TYPE "Table Row Data"
   STRUCT
      address : UInt;
      ordered : Bool;
      pbSelection : Struct
         actuate : Bool;
         animate : USInt;
      END_STRUCT;
      rtBackground : Struct
         animate : USInt;
      END_STRUCT;
      tfDropZone : Struct
         animate : USInt;
         value : WString[20];
      END_STRUCT;
      tfLine : Struct
         animate : USInt;
         value : WString[20];
      END_STRUCT;
      tfPartNumber : Struct
         animateDL : USInt;
         animateSL : USInt;
         value : WString[40];
      END_STRUCT;
      tfTime : Struct
         animate : USInt;
         value : WString[20];
      END_STRUCT;
   END_STRUCT;
END_TYPE

TYPE "Station Assignment: Button Details Data"
   STRUCT
      alloted : Struct
         animate : USInt;
         value : WString[10];
      END_STRUCT;
      critical : Struct
         animate : USInt;
         value : WString[10];
      END_STRUCT;
      label : Struct
         animate : USInt;
         value : WString[2];
      END_STRUCT;
      partNumber : Struct
         animate : USInt;
         value : WString[40];
      END_STRUCT;
      select : Struct
         actuate : Bool;
         animate : USInt;
      END_STRUCT;
   END_STRUCT;
END_TYPE

(* ===== HMI "HMI_RT_1" =====
system functions are stored by id; their names below are inferred from use
connection "HMI_Connection_2": ETHERNET, S7_1500_OMS

HMI tags "Default tag table"
   "Clock_Byte" : Byte = PLC Clock_Byte AT %MB0, 100 ms
   "HMI_screenNumber" : Int = PLC HMI.screenNumber AT %DB1.DBW0, 100 ms
   "HMI_barcode" : Barcode Screen = PLC HMI.barcode AT %DB1.DBW0, 100 ms
   "HMI_partCall_row{0}" : Table Row = PLC HMI.partCall.row[0], 100 ms
   "HMI_partCall_row{1}" : Table Row = PLC HMI.partCall.row[1], 100 ms
   "HMI_partCall_row{2}" : Table Row = PLC HMI.partCall.row[2], 100 ms
   "HMI_partCall_row{3}" : Table Row = PLC HMI.partCall.row[3], 100 ms
   "HMI_partCall_row{4}" : Table Row = PLC HMI.partCall.row[4], 100 ms
   "HMI_partCall_row{5}" : Table Row = PLC HMI.partCall.row[5], 100 ms
   "HMI_partCall_row{6}" : Table Row = PLC HMI.partCall.row[6], 100 ms
   "HMI_partCall_row{7}" : Table Row = PLC HMI.partCall.row[7], 100 ms
   "HMI_partCall_row{8}" : Table Row = PLC HMI.partCall.row[8], 100 ms
   "HMI_partCall_row{9}" : Table Row = PLC HMI.partCall.row[9], 100 ms
   "HMI_partCall_row{10}" : Table Row = PLC HMI.partCall.row[10], 100 ms
   "HMI_settings_stations_selectBtns{0}" : PB Data: Text Label = PLC HMI.settings.stations.selectBtns[0], 100 ms
   "HMI_settings_stations_selectBtns{1}" : PB Data: Text Label = PLC HMI.settings.stations.selectBtns[1], 100 ms
   "HMI_settings_stations_selectBtns{2}" : PB Data: Text Label = PLC HMI.settings.stations.selectBtns[2], 100 ms
   "HMI_settings_stations_selectBtns{3}" : PB Data: Text Label = PLC HMI.settings.stations.selectBtns[3], 100 ms
   "HMI_settings_stations_selectBtns{4}" : PB Data: Text Label = PLC HMI.settings.stations.selectBtns[4], 100 ms
   "HMI_settings_stations_selectBtns{5}" : PB Data: Text Label = PLC HMI.settings.stations.selectBtns[5], 100 ms
   "HMI_settings_stations_selectBtns{6}" : PB Data: Text Label = PLC HMI.settings.stations.selectBtns[6], 100 ms
   "HMI_settings_stations_selectBtns{7}" : PB Data: Text Label = PLC HMI.settings.stations.selectBtns[7], 100 ms
   "HMI_settings_stations_selectBtns{8}" : PB Data: Text Label = PLC HMI.settings.stations.selectBtns[8], 100 ms
   "HMI_settings_stations_selectBtns{9}" : PB Data: Text Label = PLC HMI.settings.stations.selectBtns[9], 100 ms
   "HMI_settings_stations_selectBtns{10}" : PB Data: Text Label = PLC HMI.settings.stations.selectBtns[10], 100 ms
   "HMI_settings_stations_selectBtns{11}" : PB Data: Text Label = PLC HMI.settings.stations.selectBtns[11], 100 ms
   "HMI_settings_kp8_buttons{0}" : PB Data: Text Label = PLC HMI.settings.kp8.buttons[0], 100 ms
   "HMI_settings_kp8_buttons{7}" : PB Data: Text Label = PLC HMI.settings.kp8.buttons[7], 100 ms
   "HMI_settings_kp8_buttons{3}" : PB Data: Text Label = PLC HMI.settings.kp8.buttons[3], 100 ms
   "HMI_settings_kp8_buttons{6}" : PB Data: Text Label = PLC HMI.settings.kp8.buttons[6], 100 ms
   "HMI_settings_kp8_buttons{2}" : PB Data: Text Label = PLC HMI.settings.kp8.buttons[2], 100 ms
   "HMI_settings_kp8_buttons{5}" : PB Data: Text Label = PLC HMI.settings.kp8.buttons[5], 100 ms
   "HMI_settings_kp8_buttons{1}" : PB Data: Text Label = PLC HMI.settings.kp8.buttons[1], 100 ms
   "HMI_settings_kp8_buttons{4}" : PB Data: Text Label = PLC HMI.settings.kp8.buttons[4], 100 ms
   "HMI_settings_stations_selCount" : Int = PLC HMI.settings.stations.selCount, 100 ms
   "HMI_settings_viewingStation_btns{0}" : Station Assignment: Button Details = PLC HMI.settings.viewingStation.btns[0], 100 ms
   "HMI_settings_viewingStation_btns{1}" : Station Assignment: Button Details = PLC HMI.settings.viewingStation.btns[1], 100 ms
   "HMI_settings_viewingStation_btns{2}" : Station Assignment: Button Details = PLC HMI.settings.viewingStation.btns[2], 100 ms
   "HMI_settings_viewingStation_btns{3}" : Station Assignment: Button Details = PLC HMI.settings.viewingStation.btns[3], 100 ms
   "HMI_settings_viewingStation_btns{4}" : Station Assignment: Button Details = PLC HMI.settings.viewingStation.btns[4], 100 ms
   "HMI_settings_viewingStation_btns{5}" : Station Assignment: Button Details = PLC HMI.settings.viewingStation.btns[5], 100 ms
   "HMI_settings_viewingStation_previous" : PB Data: Graphic/Text List = PLC HMI.settings.viewingStation.previous, 100 ms
   "HMI_settings_viewingStation_next" : PB Data: Graphic/Text List = PLC HMI.settings.viewingStation.next, 100 ms
   "HMI_settings_stations_selectAll" : PB Data: Text Label = PLC HMI.settings.stations.selectAll, 100 ms
   "HMI_settings_partNumber_assign" : PB Data: Text Label = PLC HMI.settings.partNumber.assign, 100 ms
   "HMI_settings_partNumber_ioField" : IO Field Data: Part Number = PLC HMI.settings.partNumber.ioField, 100 ms
   "HMI_settings_alotted_assign" : PB Data: Text Label = PLC HMI.settings.alotted.assign, 100 ms
   "HMI_settings_alotted_ioField" : IO Field Data: Timers = PLC HMI.settings.alotted.ioField, 100 ms
   "HMI_settings_critical_assign" : PB Data: Text Label = PLC HMI.settings.critical.assign, 100 ms
   "HMI_settings_critical_ioField" : IO Field Data: Timers = PLC HMI.settings.critical.ioField, 100 ms
   "HMI_settings_kp8_selectButtons" : PB Data: Text Label = PLC HMI.settings.kp8.selectButtons, 100 ms
   "HMI_settings_viewingStation_dzData" : Drop Zone Data = PLC HMI.settings.viewingStation.dzData, 100 ms
   "HMI_settings_viewingStation_lineData" : Line Label Data = PLC HMI.settings.viewingStation.lineData, 100 ms
   "HMI_settings_stations_prevGroup" : PB Data: Graphic/Text List = PLC HMI.settings.stations.prevGroup, 100 ms
   "HMI_settings_stations_nextGroup" : PB Data: Graphic/Text List = PLC HMI.settings.stations.nextGroup, 100 ms
   "HMI_settings_viewingStation_name" : WString[20] = PLC HMI.settings.viewingStation.name, 100 ms
   "HMI_tableNav_top" : PB Data: Graphic/Text List = PLC HMI.tableNav.top, 100 ms
   "HMI_tableNav_pageUp" : PB Data: Graphic/Text List = PLC HMI.tableNav.pageUp, 100 ms
   "HMI_tableNav_lineUp" : PB Data: Graphic/Text List = PLC HMI.tableNav.lineUp, 100 ms
   "HMI_tableNav_lineDown" : PB Data: Graphic/Text List = PLC HMI.tableNav.lineDown, 100 ms
   "HMI_tableNav_pageDown" : PB Data: Graphic/Text List = PLC HMI.tableNav.pageDown, 100 ms
   "HMI_tableNav_bottom" : PB Data: Graphic/Text List = PLC HMI.tableNav.bottom, 100 ms
   "HMI_simStations_stations{0}" : Station Sim Data = PLC HMI.simStations.me[0] AT %DB1.DBX0.0, 100 ms
   "HMI_simStations_me{1}" : Station Sim Data = PLC HMI.simStations.me[1], 100 ms
   "HMI_simStations_me{2}" : Station Sim Data = PLC HMI.simStations.me[2], 100 ms
   "HMI_simStations_me{3}" : Station Sim Data = PLC HMI.simStations.me[3], 100 ms
   "HMI_simStations_me{4}" : Station Sim Data = PLC HMI.simStations.me[4], 100 ms
   "HMI_simStations_me{5}" : Station Sim Data = PLC HMI.simStations.me[5], 100 ms
   "HMI_simStations_me{6}" : Station Sim Data = PLC HMI.simStations.me[6], 100 ms
   "HMI_simStations_me{7}" : Station Sim Data = PLC HMI.simStations.me[7], 100 ms
   "HMI_simStations_me{8}" : Station Sim Data = PLC HMI.simStations.me[8], 100 ms
   "HMI_simStations_me{9}" : Station Sim Data = PLC HMI.simStations.me[9], 100 ms
   "HMI_simStations_me{10}" : Station Sim Data = PLC HMI.simStations.me[10], 100 ms
   "HMI_simStations_me{11}" : Station Sim Data = PLC HMI.simStations.me[11], 100 ms
   "HMI_simStations_up" : PB Data: Graphic/Text List = PLC HMI.simStations.up, 100 ms
   "HMI_simStations_down" : PB Data: Graphic/Text List = PLC HMI.simStations.down, 100 ms
   "Log Flag" : Int = PLC "Log Buffer".logFlag AT %DB1.DBW0, 100 ms
      on ChangeValue: function_abcfba0d("Log Buffer_partReq_me{0}_address"); function_abcfba0d("Log Buffer_partReq_me{0}_timeStamp"); function_abcfba0d("Log Buffer_partReq_me{0}_reqType")
   "Log Buffer_partReq_me{0}_address" : Int = PLC "Log Buffer".partReq.me[0].address, 100 ms
   "Log Buffer_partReq_me{0}_timeStamp" : DTL = PLC "Log Buffer".partReq.me[0].timeStamp, 100 ms
   "Log Buffer_partReq_me{0}_reqType" : Int = PLC "Log Buffer".partReq.me[0].reqType, 100 ms
   "HMI_networkHealth_pnioDevices{1}" : PB Data: Text Label = PLC HMI.networkHealth.pnioDevices[1], 100 ms
   "HMI_networkHealth_pnioDevices{2}" : PB Data: Text Label = PLC HMI.networkHealth.pnioDevices[2], 1 s
   "HMI_networkHealth_pnioDevices{3}" : PB Data: Text Label = PLC HMI.networkHealth.pnioDevices[3], 1 s
   "HMI_networkHealth_pnioDevices{4}" : PB Data: Text Label = PLC HMI.networkHealth.pnioDevices[4], 1 s
   "HMI_networkHealth_pnioDevices{5}" : PB Data: Text Label = PLC HMI.networkHealth.pnioDevices[5], 1 s
   "HMI_networkHealth_pnioDevices{6}" : PB Data: Text Label = PLC HMI.networkHealth.pnioDevices[6], 1 s
   "HMI_networkHealth_pnioDevices{7}" : PB Data: Text Label = PLC HMI.networkHealth.pnioDevices[7], 1 s
   "HMI_networkHealth_pnioDevices{8}" : PB Data: Text Label = PLC HMI.networkHealth.pnioDevices[8], 1 s
   "HMI_networkHealth_pnioDevices{9}" : PB Data: Text Label = PLC HMI.networkHealth.pnioDevices[9], 1 s
   "HMI_networkHealth_pnioDevices{10}" : PB Data: Text Label = PLC HMI.networkHealth.pnioDevices[10], 1 s
   "HMI_networkHealth_pnioDevices{11}" : PB Data: Text Label = PLC HMI.networkHealth.pnioDevices[11], 1 s
   "HMI_networkHealth_pnioDevices{12}" : PB Data: Text Label = PLC HMI.networkHealth.pnioDevices[12], 1 s
   "HMI_networkHealth_pnioDevices{13}" : PB Data: Text Label = PLC HMI.networkHealth.pnioDevices[13], 1 s
   "HMI_networkHealth_pnioDevices{16}" : PB Data: Text Label = PLC HMI.networkHealth.pnioDevices[16], 1 s
   "HMI_networkHealth_pnioDevices{14}" : PB Data: Text Label = PLC HMI.networkHealth.pnioDevices[14], 1 s
   "HMI_networkHealth_pnioDevices{15}" : PB Data: Text Label = PLC HMI.networkHealth.pnioDevices[15], 1 s
   "HMI_networkHealth_pnioDevices{17}" : PB Data: Text Label = PLC HMI.networkHealth.pnioDevices[17], 1 s
   "HMI_networkHealth_pnioDevices{18}" : PB Data: Text Label = PLC HMI.networkHealth.pnioDevices[18], 1 s
   "HMI_networkHealth_pnioDevices{19}" : PB Data: Text Label = PLC HMI.networkHealth.pnioDevices[19], 1 s
   "HMI_networkHealth_pnioDevices{20}" : PB Data: Text Label = PLC HMI.networkHealth.pnioDevices[20], 1 s
   "HMI_networkHealth_pnioDevices{21}" : PB Data: Text Label = PLC HMI.networkHealth.pnioDevices[21], 1 s
   "HMI_networkHealth_pnioDevices{22}" : PB Data: Text Label = PLC HMI.networkHealth.pnioDevices[22], 1 s
   "HMI_networkHealth_pnioDevices{31}" : PB Data: Text Label = PLC HMI.networkHealth.pnioDevices[31], 1 s
   "HMI_networkHealth_pnioDevices{32}" : PB Data: Text Label = PLC HMI.networkHealth.pnioDevices[32], 1 s
   "HMI_networkHealth_pnioDevices{29}" : PB Data: Text Label = PLC HMI.networkHealth.pnioDevices[29], 1 s
   "HMI_networkHealth_pnioDevices{30}" : PB Data: Text Label = PLC HMI.networkHealth.pnioDevices[30], 1 s
   "HMI_networkHealth_pnioDevices{27}" : PB Data: Text Label = PLC HMI.networkHealth.pnioDevices[27], 1 s
   "HMI_networkHealth_pnioDevices{28}" : PB Data: Text Label = PLC HMI.networkHealth.pnioDevices[28], 1 s
   "HMI_networkHealth_pnioDevices{23}" : PB Data: Text Label = PLC HMI.networkHealth.pnioDevices[23], 1 s
   "HMI_networkHealth_pnioDevices{24}" : PB Data: Text Label = PLC HMI.networkHealth.pnioDevices[24], 1 s
   "HMI_networkHealth_pnioDevices{25}" : PB Data: Text Label = PLC HMI.networkHealth.pnioDevices[25], 1 s
   "HMI_networkHealth_pnioDevices{26}" : PB Data: Text Label = PLC HMI.networkHealth.pnioDevices[26], 1 s
   "HMI_networkHealth_pnioDevices{33}" : PB Data: Text Label = PLC HMI.networkHealth.pnioDevices[33], 1 s
   "HMI_networkHealth_pnioDevices{34}" : PB Data: Text Label = PLC HMI.networkHealth.pnioDevices[34], 1 s
   "HMI_networkHealth_pnioDevices{35}" : PB Data: Text Label = PLC HMI.networkHealth.pnioDevices[35], 1 s
   "HMI_networkHealth_pnioDevices{36}" : PB Data: Text Label = PLC HMI.networkHealth.pnioDevices[36], 1 s
   "HMI_networkHealth_pnioDevices{37}" : PB Data: Text Label = PLC HMI.networkHealth.pnioDevices[37], 1 s
   "HMI_networkHealth_pnioDevices{38}" : PB Data: Text Label = PLC HMI.networkHealth.pnioDevices[38], 1 s
   "HMI_networkHealth_pnioDevices{39}" : PB Data: Text Label = PLC HMI.networkHealth.pnioDevices[39], 1 s
   "HMI_networkHealth_pnioDevices{40}" : PB Data: Text Label = PLC HMI.networkHealth.pnioDevices[40], 1 s
   "HMI_networkHealth_pnioDevices{41}" : PB Data: Text Label = PLC HMI.networkHealth.pnioDevices[41], 1 s
   "HMI_networkHealth_pnioDevices{42}" : PB Data: Text Label = PLC HMI.networkHealth.pnioDevices[42], 1 s
   "HMI_networkHealth_pnioDevices{43}" : PB Data: Text Label = PLC HMI.networkHealth.pnioDevices[43], 1 s
   "HMI_networkHealth_pnioDevices{44}" : PB Data: Text Label = PLC HMI.networkHealth.pnioDevices[44], 1 s
   "HMI_networkHealth_pnioDevices{45}" : PB Data: Text Label = PLC HMI.networkHealth.pnioDevices[45], 1 s
   "HMI_networkHealth_pnioDevices{46}" : PB Data: Text Label = PLC HMI.networkHealth.pnioDevices[46], 1 s
   "HMI_networkHealth_pnioDevices{47}" : PB Data: Text Label = PLC HMI.networkHealth.pnioDevices[47], 1 s
   "HMI_networkHealth_pnioDevices{48}" : PB Data: Text Label = PLC HMI.networkHealth.pnioDevices[48], 1 s
   "HMI_networkHealth_et200spPopUp" : Station: ET200SP Comm Debug Data = PLC HMI.networkHealth.et200spPopUp, 1 s
   "HMI_networkHealth_kp8PopUp" : Station: KP8 Comm Debug Data = PLC HMI.networkHealth.kp8PopUp, 1 s
   "HMI_networkHealth_selectedDevice" : Int = PLC HMI.networkHealth.selectedDevice, 1 s
   "EMP IDB_stations_me{0}_partNumbers{0}" : WString[40] = PLC "EMP IDB".stations.me[0].partNumbers[0], 1 s
   "EMP IDB_stations_me{0}_partNumbers{1}" : WString[40] = PLC "EMP IDB".stations.me[0].partNumbers[1], 1 s
   "EMP IDB_stations_me{0}_partNumbers{2}" : WString[40] = PLC "EMP IDB".stations.me[0].partNumbers[2], 1 s
   "EMP IDB_stations_me{0}_partNumbers{3}" : WString[40] = PLC "EMP IDB".stations.me[0].partNumbers[3], 1 s
   "EMP IDB_stations_me{0}_partNumbers{4}" : WString[40] = PLC "EMP IDB".stations.me[0].partNumbers[4], 1 s
   "EMP IDB_stations_me{0}_partNumbers{5}" : WString[40] = PLC "EMP IDB".stations.me[0].partNumbers[5], 1 s
   "EMP IDB_stations_me{0}_partNumbers{6}" : WString[40] = PLC "EMP IDB".stations.me[0].partNumbers[6], 1 s
   "EMP IDB_stations_me{0}_partNumbers{7}" : WString[40] = PLC "EMP IDB".stations.me[0].partNumbers[7], 1 s
   "EMP IDB_stations_me{1}_partNumbers{0}" : WString[40] = PLC "EMP IDB".stations.me[1].partNumbers[0], 1 s
   "EMP IDB_stations_me{1}_partNumbers{1}" : WString[40] = PLC "EMP IDB".stations.me[1].partNumbers[1], 1 s
   "EMP IDB_stations_me{1}_partNumbers{2}" : WString[40] = PLC "EMP IDB".stations.me[1].partNumbers[2], 1 s
   "EMP IDB_stations_me{1}_partNumbers{3}" : WString[40] = PLC "EMP IDB".stations.me[1].partNumbers[3], 1 s
   "EMP IDB_stations_me{1}_partNumbers{4}" : WString[40] = PLC "EMP IDB".stations.me[1].partNumbers[4], 1 s
   "EMP IDB_stations_me{1}_partNumbers{5}" : WString[40] = PLC "EMP IDB".stations.me[1].partNumbers[5], 1 s
   "EMP IDB_stations_me{1}_partNumbers{6}" : WString[40] = PLC "EMP IDB".stations.me[1].partNumbers[6], 1 s
   "EMP IDB_stations_me{1}_partNumbers{7}" : WString[40] = PLC "EMP IDB".stations.me[1].partNumbers[7], 1 s
   "EMP IDB_stations_me{2}_partNumbers{0}" : WString[40] = PLC "EMP IDB".stations.me[2].partNumbers[0], 1 s
   "EMP IDB_stations_me{2}_partNumbers{1}" : WString[40] = PLC "EMP IDB".stations.me[2].partNumbers[1], 1 s
   "EMP IDB_stations_me{2}_partNumbers{2}" : WString[40] = PLC "EMP IDB".stations.me[2].partNumbers[2], 1 s
   "EMP IDB_stations_me{2}_partNumbers{3}" : WString[40] = PLC "EMP IDB".stations.me[2].partNumbers[3], 1 s
   "EMP IDB_stations_me{2}_partNumbers{4}" : WString[40] = PLC "EMP IDB".stations.me[2].partNumbers[4], 1 s
   "EMP IDB_stations_me{2}_partNumbers{5}" : WString[40] = PLC "EMP IDB".stations.me[2].partNumbers[5], 1 s
   "EMP IDB_stations_me{2}_partNumbers{6}" : WString[40] = PLC "EMP IDB".stations.me[2].partNumbers[6], 1 s
   "EMP IDB_stations_me{2}_partNumbers{7}" : WString[40] = PLC "EMP IDB".stations.me[2].partNumbers[7], 1 s
   "EMP IDB_stations_me{3}_partOrdered{0}" : Bool = PLC "EMP IDB".stations.me[3].partOrdered[0], 1 s
   "EMP IDB_stations_me{3}_partOrdered{1}" : Bool = PLC "EMP IDB".stations.me[3].partOrdered[1], 1 s
   "EMP IDB_stations_me{3}_partOrdered{2}" : Bool = PLC "EMP IDB".stations.me[3].partOrdered[2], 1 s
   "EMP IDB_stations_me{3}_partOrdered{3}" : Bool = PLC "EMP IDB".stations.me[3].partOrdered[3], 1 s
   "EMP IDB_stations_me{3}_partOrdered{4}" : Bool = PLC "EMP IDB".stations.me[3].partOrdered[4], 1 s
   "EMP IDB_stations_me{3}_partOrdered{5}" : Bool = PLC "EMP IDB".stations.me[3].partOrdered[5], 1 s
   "EMP IDB_stations_me{3}_partOrdered{6}" : Bool = PLC "EMP IDB".stations.me[3].partOrdered[6], 1 s
   "EMP IDB_stations_me{3}_partOrdered{7}" : Bool = PLC "EMP IDB".stations.me[3].partOrdered[7], 1 s
   "EMP IDB_stations_me{4}_partNumbers{0}" : WString[40] = PLC "EMP IDB".stations.me[4].partNumbers[0], 1 s
   "EMP IDB_stations_me{4}_partNumbers{1}" : WString[40] = PLC "EMP IDB".stations.me[4].partNumbers[1], 1 s
   "EMP IDB_stations_me{4}_partNumbers{2}" : WString[40] = PLC "EMP IDB".stations.me[4].partNumbers[2], 1 s
   "EMP IDB_stations_me{4}_partNumbers{3}" : WString[40] = PLC "EMP IDB".stations.me[4].partNumbers[3], 1 s
   "EMP IDB_stations_me{4}_partNumbers{4}" : WString[40] = PLC "EMP IDB".stations.me[4].partNumbers[4], 1 s
   "EMP IDB_stations_me{4}_partNumbers{5}" : WString[40] = PLC "EMP IDB".stations.me[4].partNumbers[5], 1 s
   "EMP IDB_stations_me{4}_partNumbers{6}" : WString[40] = PLC "EMP IDB".stations.me[4].partNumbers[6], 1 s
   "EMP IDB_stations_me{4}_partNumbers{7}" : WString[40] = PLC "EMP IDB".stations.me[4].partNumbers[7], 1 s
   "EMP IDB_stations_me{5}_partNumbers{0}" : WString[40] = PLC "EMP IDB".stations.me[5].partNumbers[0], 1 s
   "EMP IDB_stations_me{5}_partNumbers{1}" : WString[40] = PLC "EMP IDB".stations.me[5].partNumbers[1], 1 s
   "EMP IDB_stations_me{5}_partNumbers{2}" : WString[40] = PLC "EMP IDB".stations.me[5].partNumbers[2], 1 s
   "EMP IDB_stations_me{5}_partNumbers{3}" : WString[40] = PLC "EMP IDB".stations.me[5].partNumbers[3], 1 s
   "EMP IDB_stations_me{5}_partNumbers{4}" : WString[40] = PLC "EMP IDB".stations.me[5].partNumbers[4], 1 s
   "EMP IDB_stations_me{5}_partNumbers{5}" : WString[40] = PLC "EMP IDB".stations.me[5].partNumbers[5], 1 s
   "EMP IDB_stations_me{5}_partNumbers{6}" : WString[40] = PLC "EMP IDB".stations.me[5].partNumbers[6], 1 s
   "EMP IDB_stations_me{5}_partNumbers{7}" : WString[40] = PLC "EMP IDB".stations.me[5].partNumbers[7], 1 s
   "EMP IDB_stations_me{6}_partNumbers{0}" : WString[40] = PLC "EMP IDB".stations.me[6].partNumbers[0], 1 s
   "EMP IDB_stations_me{6}_partNumbers{1}" : WString[40] = PLC "EMP IDB".stations.me[6].partNumbers[1], 1 s
   "EMP IDB_stations_me{6}_partNumbers{2}" : WString[40] = PLC "EMP IDB".stations.me[6].partNumbers[2], 1 s
   "EMP IDB_stations_me{6}_partNumbers{3}" : WString[40] = PLC "EMP IDB".stations.me[6].partNumbers[3], 1 s
   "EMP IDB_stations_me{6}_partNumbers{4}" : WString[40] = PLC "EMP IDB".stations.me[6].partNumbers[4], 1 s
   "EMP IDB_stations_me{6}_partNumbers{5}" : WString[40] = PLC "EMP IDB".stations.me[6].partNumbers[5], 1 s
   "EMP IDB_stations_me{6}_partNumbers{6}" : WString[40] = PLC "EMP IDB".stations.me[6].partNumbers[6], 1 s
   "EMP IDB_stations_me{6}_partNumbers{7}" : WString[40] = PLC "EMP IDB".stations.me[6].partNumbers[7], 1 s
   "EMP IDB_stations_me{7}_partNumbers{0}" : WString[40] = PLC "EMP IDB".stations.me[7].partNumbers[0], 1 s
   "EMP IDB_stations_me{7}_partNumbers{1}" : WString[40] = PLC "EMP IDB".stations.me[7].partNumbers[1], 1 s
   "EMP IDB_stations_me{7}_partNumbers{2}" : WString[40] = PLC "EMP IDB".stations.me[7].partNumbers[2], 1 s
   "EMP IDB_stations_me{7}_partNumbers{3}" : WString[40] = PLC "EMP IDB".stations.me[7].partNumbers[3], 1 s
   "EMP IDB_stations_me{7}_partNumbers{4}" : WString[40] = PLC "EMP IDB".stations.me[7].partNumbers[4], 1 s
   "EMP IDB_stations_me{7}_partNumbers{5}" : WString[40] = PLC "EMP IDB".stations.me[7].partNumbers[5], 1 s
   "EMP IDB_stations_me{7}_partNumbers{6}" : WString[40] = PLC "EMP IDB".stations.me[7].partNumbers[6], 1 s
   "EMP IDB_stations_me{7}_partNumbers{7}" : WString[40] = PLC "EMP IDB".stations.me[7].partNumbers[7], 1 s
   "EMP IDB_stations_me{8}_partNumbers{0}" : WString[40] = PLC "EMP IDB".stations.me[8].partNumbers[0], 1 s
   "EMP IDB_stations_me{8}_partNumbers{1}" : WString[40] = PLC "EMP IDB".stations.me[8].partNumbers[1], 1 s
   "EMP IDB_stations_me{8}_partNumbers{2}" : WString[40] = PLC "EMP IDB".stations.me[8].partNumbers[2], 1 s
   "EMP IDB_stations_me{8}_partNumbers{3}" : WString[40] = PLC "EMP IDB".stations.me[8].partNumbers[3], 1 s
   "EMP IDB_stations_me{8}_partNumbers{4}" : WString[40] = PLC "EMP IDB".stations.me[8].partNumbers[4], 1 s
   "EMP IDB_stations_me{8}_partNumbers{5}" : WString[40] = PLC "EMP IDB".stations.me[8].partNumbers[5], 1 s
   "EMP IDB_stations_me{8}_partNumbers{6}" : WString[40] = PLC "EMP IDB".stations.me[8].partNumbers[6], 1 s
   "EMP IDB_stations_me{8}_partNumbers{7}" : WString[40] = PLC "EMP IDB".stations.me[8].partNumbers[7], 1 s
   "EMP IDB_stations_me{9}_partNumbers{0}" : WString[40] = PLC "EMP IDB".stations.me[9].partNumbers[0], 1 s
   "EMP IDB_stations_me{9}_partNumbers{1}" : WString[40] = PLC "EMP IDB".stations.me[9].partNumbers[1], 1 s
   "EMP IDB_stations_me{9}_partNumbers{2}" : WString[40] = PLC "EMP IDB".stations.me[9].partNumbers[2], 1 s
   "EMP IDB_stations_me{9}_partNumbers{3}" : WString[40] = PLC "EMP IDB".stations.me[9].partNumbers[3], 1 s
   "EMP IDB_stations_me{9}_partNumbers{4}" : WString[40] = PLC "EMP IDB".stations.me[9].partNumbers[4], 1 s
   "EMP IDB_stations_me{9}_partNumbers{5}" : WString[40] = PLC "EMP IDB".stations.me[9].partNumbers[5], 1 s
   "EMP IDB_stations_me{9}_partNumbers{6}" : WString[40] = PLC "EMP IDB".stations.me[9].partNumbers[6], 1 s
   "EMP IDB_stations_me{9}_partNumbers{7}" : WString[40] = PLC "EMP IDB".stations.me[9].partNumbers[7], 1 s
   "EMP IDB_stations_me{10}_partNumbers{0}" : WString[40] = PLC "EMP IDB".stations.me[10].partNumbers[0], 1 s
   "EMP IDB_stations_me{10}_partNumbers{1}" : WString[40] = PLC "EMP IDB".stations.me[10].partNumbers[1], 1 s
   "EMP IDB_stations_me{10}_partNumbers{2}" : WString[40] = PLC "EMP IDB".stations.me[10].partNumbers[2], 1 s
   "EMP IDB_stations_me{10}_partNumbers{3}" : WString[40] = PLC "EMP IDB".stations.me[10].partNumbers[3], 1 s
   "EMP IDB_stations_me{10}_partNumbers{4}" : WString[40] = PLC "EMP IDB".stations.me[10].partNumbers[4], 1 s
   "EMP IDB_stations_me{10}_partNumbers{5}" : WString[40] = PLC "EMP IDB".stations.me[10].partNumbers[5], 1 s
   "EMP IDB_stations_me{10}_partNumbers{6}" : WString[40] = PLC "EMP IDB".stations.me[10].partNumbers[6], 1 s
   "EMP IDB_stations_me{10}_partNumbers{7}" : WString[40] = PLC "EMP IDB".stations.me[10].partNumbers[7], 1 s
   "EMP IDB_stations_me{11}_partNumbers{0}" : WString[40] = PLC "EMP IDB".stations.me[11].partNumbers[0], 1 s
   "EMP IDB_stations_me{11}_partNumbers{1}" : WString[40] = PLC "EMP IDB".stations.me[11].partNumbers[1], 1 s
   "EMP IDB_stations_me{11}_partNumbers{2}" : WString[40] = PLC "EMP IDB".stations.me[11].partNumbers[2], 1 s
   "EMP IDB_stations_me{11}_partNumbers{3}" : WString[40] = PLC "EMP IDB".stations.me[11].partNumbers[3], 1 s
   "EMP IDB_stations_me{11}_partNumbers{4}" : WString[40] = PLC "EMP IDB".stations.me[11].partNumbers[4], 1 s
   "EMP IDB_stations_me{11}_partNumbers{5}" : WString[40] = PLC "EMP IDB".stations.me[11].partNumbers[5], 1 s
   "EMP IDB_stations_me{11}_partNumbers{6}" : WString[40] = PLC "EMP IDB".stations.me[11].partNumbers[6], 1 s
   "EMP IDB_stations_me{11}_partNumbers{7}" : WString[40] = PLC "EMP IDB".stations.me[11].partNumbers[7], 1 s
   "EMP IDB_stations_me{12}_partNumbers{0}" : WString[40] = PLC "EMP IDB".stations.me[12].partNumbers[0], 1 s
   "EMP IDB_stations_me{12}_partNumbers{1}" : WString[40] = PLC "EMP IDB".stations.me[12].partNumbers[1], 1 s
   "EMP IDB_stations_me{12}_partNumbers{2}" : WString[40] = PLC "EMP IDB".stations.me[12].partNumbers[2], 1 s
   "EMP IDB_stations_me{12}_partNumbers{3}" : WString[40] = PLC "EMP IDB".stations.me[12].partNumbers[3], 1 s
   "EMP IDB_stations_me{12}_partNumbers{4}" : WString[40] = PLC "EMP IDB".stations.me[12].partNumbers[4], 1 s
   "EMP IDB_stations_me{12}_partNumbers{5}" : WString[40] = PLC "EMP IDB".stations.me[12].partNumbers[5], 1 s
   "EMP IDB_stations_me{12}_partNumbers{6}" : WString[40] = PLC "EMP IDB".stations.me[12].partNumbers[6], 1 s
   "EMP IDB_stations_me{12}_partNumbers{7}" : WString[40] = PLC "EMP IDB".stations.me[12].partNumbers[7], 1 s
   "EMP IDB_stations_me{13}_partNumbers{0}" : WString[40] = PLC "EMP IDB".stations.me[13].partNumbers[0], 1 s
   "EMP IDB_stations_me{13}_partNumbers{1}" : WString[40] = PLC "EMP IDB".stations.me[13].partNumbers[1], 1 s
   "EMP IDB_stations_me{13}_partNumbers{2}" : WString[40] = PLC "EMP IDB".stations.me[13].partNumbers[2], 1 s
   "EMP IDB_stations_me{13}_partNumbers{3}" : WString[40] = PLC "EMP IDB".stations.me[13].partNumbers[3], 1 s
   "EMP IDB_stations_me{13}_partNumbers{4}" : WString[40] = PLC "EMP IDB".stations.me[13].partNumbers[4], 1 s
   "EMP IDB_stations_me{13}_partNumbers{5}" : WString[40] = PLC "EMP IDB".stations.me[13].partNumbers[5], 1 s
   "EMP IDB_stations_me{13}_partNumbers{6}" : WString[40] = PLC "EMP IDB".stations.me[13].partNumbers[6], 1 s
   "EMP IDB_stations_me{13}_partNumbers{7}" : WString[40] = PLC "EMP IDB".stations.me[13].partNumbers[7], 1 s
   "EMP IDB_stations_me{14}_partNumbers{0}" : WString[40] = PLC "EMP IDB".stations.me[14].partNumbers[0], 1 s
   "EMP IDB_stations_me{14}_partNumbers{1}" : WString[40] = PLC "EMP IDB".stations.me[14].partNumbers[1], 1 s
   "EMP IDB_stations_me{14}_partNumbers{2}" : WString[40] = PLC "EMP IDB".stations.me[14].partNumbers[2], 1 s
   "EMP IDB_stations_me{14}_partNumbers{3}" : WString[40] = PLC "EMP IDB".stations.me[14].partNumbers[3], 1 s
   "EMP IDB_stations_me{14}_partNumbers{4}" : WString[40] = PLC "EMP IDB".stations.me[14].partNumbers[4], 1 s
   "EMP IDB_stations_me{14}_partNumbers{5}" : WString[40] = PLC "EMP IDB".stations.me[14].partNumbers[5], 1 s
   "EMP IDB_stations_me{14}_partNumbers{6}" : WString[40] = PLC "EMP IDB".stations.me[14].partNumbers[6], 1 s
   "EMP IDB_stations_me{14}_partNumbers{7}" : WString[40] = PLC "EMP IDB".stations.me[14].partNumbers[7], 1 s
   "EMP IDB_stations_me{15}_partNumbers{0}" : WString[40] = PLC "EMP IDB".stations.me[15].partNumbers[0], 1 s
   "EMP IDB_stations_me{15}_partNumbers{1}" : WString[40] = PLC "EMP IDB".stations.me[15].partNumbers[1], 1 s
   "EMP IDB_stations_me{15}_partNumbers{2}" : WString[40] = PLC "EMP IDB".stations.me[15].partNumbers[2], 1 s
   "EMP IDB_stations_me{15}_partNumbers{3}" : WString[40] = PLC "EMP IDB".stations.me[15].partNumbers[3], 1 s
   "EMP IDB_stations_me{15}_partNumbers{4}" : WString[40] = PLC "EMP IDB".stations.me[15].partNumbers[4], 1 s
   "EMP IDB_stations_me{15}_partNumbers{5}" : WString[40] = PLC "EMP IDB".stations.me[15].partNumbers[5], 1 s
   "EMP IDB_stations_me{15}_partNumbers{6}" : WString[40] = PLC "EMP IDB".stations.me[15].partNumbers[6], 1 s
   "EMP IDB_stations_me{15}_partNumbers{7}" : WString[40] = PLC "EMP IDB".stations.me[15].partNumbers[7], 1 s
   "EMP IDB_stations_me{16}_partNumbers{0}" : WString[40] = PLC "EMP IDB".stations.me[16].partNumbers[0], 1 s
   "EMP IDB_stations_me{16}_partNumbers{1}" : WString[40] = PLC "EMP IDB".stations.me[16].partNumbers[1], 1 s
   "EMP IDB_stations_me{16}_partNumbers{2}" : WString[40] = PLC "EMP IDB".stations.me[16].partNumbers[2], 1 s
   "EMP IDB_stations_me{16}_partNumbers{3}" : WString[40] = PLC "EMP IDB".stations.me[16].partNumbers[3], 1 s
   "EMP IDB_stations_me{16}_partNumbers{4}" : WString[40] = PLC "EMP IDB".stations.me[16].partNumbers[4], 1 s
   "EMP IDB_stations_me{16}_partNumbers{5}" : WString[40] = PLC "EMP IDB".stations.me[16].partNumbers[5], 1 s
   "EMP IDB_stations_me{16}_partNumbers{6}" : WString[40] = PLC "EMP IDB".stations.me[16].partNumbers[6], 1 s
   "EMP IDB_stations_me{16}_partNumbers{7}" : WString[40] = PLC "EMP IDB".stations.me[16].partNumbers[7], 1 s
   "EMP IDB_stations_me{17}_partNumbers{0}" : WString[40] = PLC "EMP IDB".stations.me[17].partNumbers[0], 1 s
   "EMP IDB_stations_me{17}_partNumbers{1}" : WString[40] = PLC "EMP IDB".stations.me[17].partNumbers[1], 1 s
   "EMP IDB_stations_me{17}_partNumbers{2}" : WString[40] = PLC "EMP IDB".stations.me[17].partNumbers[2], 1 s
   "EMP IDB_stations_me{17}_partNumbers{3}" : WString[40] = PLC "EMP IDB".stations.me[17].partNumbers[3], 1 s
   "EMP IDB_stations_me{17}_partNumbers{4}" : WString[40] = PLC "EMP IDB".stations.me[17].partNumbers[4], 1 s
   "EMP IDB_stations_me{17}_partNumbers{5}" : WString[40] = PLC "EMP IDB".stations.me[17].partNumbers[5], 1 s
   "EMP IDB_stations_me{17}_partNumbers{6}" : WString[40] = PLC "EMP IDB".stations.me[17].partNumbers[6], 1 s
   "EMP IDB_stations_me{17}_partNumbers{7}" : WString[40] = PLC "EMP IDB".stations.me[17].partNumbers[7], 1 s
   "EMP IDB_stations_me{18}_partNumbers{0}" : WString[40] = PLC "EMP IDB".stations.me[18].partNumbers[0], 1 s
   "EMP IDB_stations_me{18}_partNumbers{1}" : WString[40] = PLC "EMP IDB".stations.me[18].partNumbers[1], 1 s
   "EMP IDB_stations_me{18}_partNumbers{2}" : WString[40] = PLC "EMP IDB".stations.me[18].partNumbers[2], 1 s
   "EMP IDB_stations_me{18}_partNumbers{3}" : WString[40] = PLC "EMP IDB".stations.me[18].partNumbers[3], 1 s
   "EMP IDB_stations_me{18}_partNumbers{4}" : WString[40] = PLC "EMP IDB".stations.me[18].partNumbers[4], 1 s
   "EMP IDB_stations_me{18}_partNumbers{5}" : WString[40] = PLC "EMP IDB".stations.me[18].partNumbers[5], 1 s
   "EMP IDB_stations_me{18}_partNumbers{6}" : WString[40] = PLC "EMP IDB".stations.me[18].partNumbers[6], 1 s
   "EMP IDB_stations_me{18}_partNumbers{7}" : WString[40] = PLC "EMP IDB".stations.me[18].partNumbers[7], 1 s
   "EMP IDB_stations_me{19}_partNumbers{0}" : WString[40] = PLC "EMP IDB".stations.me[19].partNumbers[0], 1 s
   "EMP IDB_stations_me{19}_partNumbers{1}" : WString[40] = PLC "EMP IDB".stations.me[19].partNumbers[1], 1 s
   "EMP IDB_stations_me{19}_partNumbers{2}" : WString[40] = PLC "EMP IDB".stations.me[19].partNumbers[2], 1 s
   "EMP IDB_stations_me{19}_partNumbers{3}" : WString[40] = PLC "EMP IDB".stations.me[19].partNumbers[3], 1 s
   "EMP IDB_stations_me{19}_partNumbers{4}" : WString[40] = PLC "EMP IDB".stations.me[19].partNumbers[4], 1 s
   "EMP IDB_stations_me{19}_partNumbers{5}" : WString[40] = PLC "EMP IDB".stations.me[19].partNumbers[5], 1 s
   "EMP IDB_stations_me{19}_partNumbers{6}" : WString[40] = PLC "EMP IDB".stations.me[19].partNumbers[6], 1 s
   "EMP IDB_stations_me{19}_partNumbers{7}" : WString[40] = PLC "EMP IDB".stations.me[19].partNumbers[7], 1 s
   "EMP IDB_stations_me{20}_partNumbers{0}" : WString[40] = PLC "EMP IDB".stations.me[20].partNumbers[0], 1 s
   "EMP IDB_stations_me{20}_partNumbers{1}" : WString[40] = PLC "EMP IDB".stations.me[20].partNumbers[1], 1 s
   "EMP IDB_stations_me{20}_partNumbers{2}" : WString[40] = PLC "EMP IDB".stations.me[20].partNumbers[2], 1 s
   "EMP IDB_stations_me{20}_partNumbers{3}" : WString[40] = PLC "EMP IDB".stations.me[20].partNumbers[3], 1 s
   "EMP IDB_stations_me{20}_partNumbers{4}" : WString[40] = PLC "EMP IDB".stations.me[20].partNumbers[4], 1 s
   "EMP IDB_stations_me{20}_partNumbers{5}" : WString[40] = PLC "EMP IDB".stations.me[20].partNumbers[5], 1 s
   "EMP IDB_stations_me{20}_partNumbers{6}" : WString[40] = PLC "EMP IDB".stations.me[20].partNumbers[6], 1 s
   "EMP IDB_stations_me{20}_partNumbers{7}" : WString[40] = PLC "EMP IDB".stations.me[20].partNumbers[7], 1 s
   "EMP IDB_stations_me{21}_partNumbers{0}" : WString[40] = PLC "EMP IDB".stations.me[21].partNumbers[0], 1 s
   "EMP IDB_stations_me{21}_partNumbers{1}" : WString[40] = PLC "EMP IDB".stations.me[21].partNumbers[1], 1 s
   "EMP IDB_stations_me{21}_partNumbers{2}" : WString[40] = PLC "EMP IDB".stations.me[21].partNumbers[2], 1 s
   "EMP IDB_stations_me{21}_partNumbers{3}" : WString[40] = PLC "EMP IDB".stations.me[21].partNumbers[3], 1 s
   "EMP IDB_stations_me{21}_partNumbers{4}" : WString[40] = PLC "EMP IDB".stations.me[21].partNumbers[4], 1 s
   "EMP IDB_stations_me{21}_partNumbers{5}" : WString[40] = PLC "EMP IDB".stations.me[21].partNumbers[5], 1 s
   "EMP IDB_stations_me{21}_partNumbers{6}" : WString[40] = PLC "EMP IDB".stations.me[21].partNumbers[6], 1 s
   "EMP IDB_stations_me{21}_partNumbers{7}" : WString[40] = PLC "EMP IDB".stations.me[21].partNumbers[7], 1 s
   "EMP IDB_stations_me{22}_partNumbers{0}" : WString[40] = PLC "EMP IDB".stations.me[22].partNumbers[0], 1 s
   "EMP IDB_stations_me{22}_partNumbers{1}" : WString[40] = PLC "EMP IDB".stations.me[22].partNumbers[1], 1 s
   "EMP IDB_stations_me{22}_partNumbers{2}" : WString[40] = PLC "EMP IDB".stations.me[22].partNumbers[2], 1 s
   "EMP IDB_stations_me{22}_partNumbers{3}" : WString[40] = PLC "EMP IDB".stations.me[22].partNumbers[3], 1 s
   "EMP IDB_stations_me{22}_partNumbers{4}" : WString[40] = PLC "EMP IDB".stations.me[22].partNumbers[4], 1 s
   "EMP IDB_stations_me{22}_partNumbers{5}" : WString[40] = PLC "EMP IDB".stations.me[22].partNumbers[5], 1 s
   "EMP IDB_stations_me{22}_partNumbers{6}" : WString[40] = PLC "EMP IDB".stations.me[22].partNumbers[6], 1 s
   "EMP IDB_stations_me{22}_partNumbers{7}" : WString[40] = PLC "EMP IDB".stations.me[22].partNumbers[7], 1 s
   "EMP IDB_stations_me{23}_partNumbers{0}" : WString[40] = PLC "EMP IDB".stations.me[23].partNumbers[0], 1 s
   "EMP IDB_stations_me{23}_partNumbers{1}" : WString[40] = PLC "EMP IDB".stations.me[23].partNumbers[1], 1 s
   "EMP IDB_stations_me{23}_partNumbers{2}" : WString[40] = PLC "EMP IDB".stations.me[23].partNumbers[2], 1 s
   "EMP IDB_stations_me{23}_partNumbers{3}" : WString[40] = PLC "EMP IDB".stations.me[23].partNumbers[3], 1 s
   "EMP IDB_stations_me{23}_partNumbers{4}" : WString[40] = PLC "EMP IDB".stations.me[23].partNumbers[4], 1 s
   "EMP IDB_stations_me{23}_partNumbers{5}" : WString[40] = PLC "EMP IDB".stations.me[23].partNumbers[5], 1 s
   "EMP IDB_stations_me{23}_partNumbers{6}" : WString[40] = PLC "EMP IDB".stations.me[23].partNumbers[6], 1 s
   "EMP IDB_stations_me{23}_partNumbers{7}" : WString[40] = PLC "EMP IDB".stations.me[23].partNumbers[7], 1 s
   "EMP IDB_stations_me{3}_partNumbers{0}" : WString[40] = PLC "EMP IDB".stations.me[3].partNumbers[0], 1 s

text list "Station Selection Single": 0 'Select a Station to View'; 1 'Assignments'

recipe "VOLVO 16 01": Button 0 <- "EMP IDB_stations_me{0}_partNumbers{0}", Button 1 <- "EMP IDB_stations_me{0}_partNumbers{1}", Button 2 <- "EMP IDB_stations_me{0}_partNumbers{2}", Button 3 <- "EMP IDB_stations_me{0}_partNumbers{3}", Button 4 <- "EMP IDB_stations_me{0}_partNumbers{4}", Button 5 <- "EMP IDB_stations_me{0}_partNumbers{5}", Button 6 <- "EMP IDB_stations_me{0}_partNumbers{6}", Button 7 <- "EMP IDB_stations_me{0}_partNumbers{7}"

recipe "VOLVO 16 02": Button 0 <- "EMP IDB_stations_me{1}_partNumbers{0}", Button 1 <- "EMP IDB_stations_me{1}_partNumbers{1}", Button 2 <- "EMP IDB_stations_me{1}_partNumbers{2}", Button 3 <- "EMP IDB_stations_me{1}_partNumbers{3}", Button 4 <- "EMP IDB_stations_me{1}_partNumbers{4}", Button 5 <- "EMP IDB_stations_me{1}_partNumbers{5}", Button 6 <- "EMP IDB_stations_me{1}_partNumbers{6}", Button 7 <- "EMP IDB_stations_me{1}_partNumbers{7}"

recipe "VOLVO 16 03": Button 0 <- "EMP IDB_stations_me{2}_partNumbers{0}", Button 1 <- "EMP IDB_stations_me{2}_partNumbers{1}", Button 2 <- "EMP IDB_stations_me{2}_partNumbers{2}", Button 3 <- "EMP IDB_stations_me{2}_partNumbers{3}", Button 4 <- "EMP IDB_stations_me{2}_partNumbers{4}", Button 5 <- "EMP IDB_stations_me{2}_partNumbers{5}", Button 6 <- "EMP IDB_stations_me{2}_partNumbers{6}", Button 7 <- "EMP IDB_stations_me{2}_partNumbers{7}"

recipe "VOLVO 16 04": Button 0 <- "EMP IDB_stations_me{3}_partNumbers{0}", Button 1, Button 2, Button 3, Button 4, Button 5, Button 6, Button 7, Recipe_element_1

recipe "VOLVO 16 05": Button 0 <- "EMP IDB_stations_me{4}_partNumbers{0}", Button 1 <- "EMP IDB_stations_me{4}_partNumbers{1}", Button 2 <- "EMP IDB_stations_me{4}_partNumbers{2}", Button 3 <- "EMP IDB_stations_me{4}_partNumbers{3}", Button 4 <- "EMP IDB_stations_me{4}_partNumbers{4}", Button 5 <- "EMP IDB_stations_me{4}_partNumbers{5}", Button 6 <- "EMP IDB_stations_me{4}_partNumbers{6}", Button 7 <- "EMP IDB_stations_me{4}_partNumbers{7}"

recipe "VOLVO 16 06": Button 0 <- "EMP IDB_stations_me{5}_partNumbers{0}", Button 1 <- "EMP IDB_stations_me{5}_partNumbers{1}", Button 2 <- "EMP IDB_stations_me{5}_partNumbers{2}", Button 3 <- "EMP IDB_stations_me{5}_partNumbers{3}", Button 4 <- "EMP IDB_stations_me{5}_partNumbers{4}", Button 5 <- "EMP IDB_stations_me{5}_partNumbers{5}", Button 6 <- "EMP IDB_stations_me{5}_partNumbers{6}", Button 7 <- "EMP IDB_stations_me{5}_partNumbers{7}"

recipe "VOLVO 16 07": Button 0 <- "EMP IDB_stations_me{6}_partNumbers{0}", Button 1 <- "EMP IDB_stations_me{6}_partNumbers{1}", Button 2 <- "EMP IDB_stations_me{6}_partNumbers{2}", Button 3 <- "EMP IDB_stations_me{6}_partNumbers{3}", Button 4 <- "EMP IDB_stations_me{6}_partNumbers{4}", Button 5 <- "EMP IDB_stations_me{6}_partNumbers{5}", Button 6 <- "EMP IDB_stations_me{6}_partNumbers{6}", Button 7 <- "EMP IDB_stations_me{6}_partNumbers{7}"

recipe "VOLVO 16 08": Button 0 <- "EMP IDB_stations_me{7}_partNumbers{0}", Button 1 <- "EMP IDB_stations_me{7}_partNumbers{1}", Button 2 <- "EMP IDB_stations_me{7}_partNumbers{2}", Button 3 <- "EMP IDB_stations_me{7}_partNumbers{3}", Button 4 <- "EMP IDB_stations_me{7}_partNumbers{4}", Button 5 <- "EMP IDB_stations_me{7}_partNumbers{5}", Button 6 <- "EMP IDB_stations_me{7}_partNumbers{6}", Button 7 <- "EMP IDB_stations_me{7}_partNumbers{7}"

recipe "VOLVO 16 09": Button 0 <- "EMP IDB_stations_me{8}_partNumbers{0}", Button 1 <- "EMP IDB_stations_me{8}_partNumbers{1}", Button 2 <- "EMP IDB_stations_me{8}_partNumbers{2}", Button 3 <- "EMP IDB_stations_me{8}_partNumbers{3}", Button 4 <- "EMP IDB_stations_me{8}_partNumbers{4}", Button 5 <- "EMP IDB_stations_me{8}_partNumbers{5}", Button 6 <- "EMP IDB_stations_me{8}_partNumbers{6}", Button 7 <- "EMP IDB_stations_me{8}_partNumbers{7}"

recipe "VOLVO 16 10": Button 0 <- "EMP IDB_stations_me{9}_partNumbers{0}", Button 1 <- "EMP IDB_stations_me{9}_partNumbers{1}", Button 2 <- "EMP IDB_stations_me{9}_partNumbers{2}", Button 3 <- "EMP IDB_stations_me{9}_partNumbers{3}", Button 4 <- "EMP IDB_stations_me{9}_partNumbers{4}", Button 5 <- "EMP IDB_stations_me{9}_partNumbers{5}", Button 6 <- "EMP IDB_stations_me{9}_partNumbers{6}", Button 7 <- "EMP IDB_stations_me{9}_partNumbers{7}"

recipe "VOLVO 16 11": Button 0 <- "EMP IDB_stations_me{10}_partNumbers{0}", Button 1 <- "EMP IDB_stations_me{10}_partNumbers{1}", Button 2 <- "EMP IDB_stations_me{10}_partNumbers{2}", Button 3 <- "EMP IDB_stations_me{10}_partNumbers{3}", Button 4 <- "EMP IDB_stations_me{10}_partNumbers{4}", Button 5 <- "EMP IDB_stations_me{10}_partNumbers{5}", Button 6 <- "EMP IDB_stations_me{10}_partNumbers{6}", Button 7 <- "EMP IDB_stations_me{10}_partNumbers{7}"

recipe "CHM 01": Button 0 <- "EMP IDB_stations_me{11}_partNumbers{0}", Button 1 <- "EMP IDB_stations_me{11}_partNumbers{1}", Button 2 <- "EMP IDB_stations_me{11}_partNumbers{2}", Button 3 <- "EMP IDB_stations_me{11}_partNumbers{3}", Button 4 <- "EMP IDB_stations_me{11}_partNumbers{4}", Button 5 <- "EMP IDB_stations_me{11}_partNumbers{5}", Button 6 <- "EMP IDB_stations_me{11}_partNumbers{6}", Button 7 <- "EMP IDB_stations_me{11}_partNumbers{7}"

recipe "CHM 02": Button 0 <- "EMP IDB_stations_me{12}_partNumbers{0}", Button 1 <- "EMP IDB_stations_me{12}_partNumbers{1}", Button 2 <- "EMP IDB_stations_me{12}_partNumbers{2}", Button 3 <- "EMP IDB_stations_me{12}_partNumbers{3}", Button 4 <- "EMP IDB_stations_me{12}_partNumbers{4}", Button 5 <- "EMP IDB_stations_me{12}_partNumbers{5}", Button 6 <- "EMP IDB_stations_me{12}_partNumbers{6}", Button 7 <- "EMP IDB_stations_me{12}_partNumbers{7}"

recipe "CHM 03": Button 0 <- "EMP IDB_stations_me{13}_partNumbers{0}", Button 1 <- "EMP IDB_stations_me{13}_partNumbers{1}", Button 2 <- "EMP IDB_stations_me{13}_partNumbers{2}", Button 3 <- "EMP IDB_stations_me{13}_partNumbers{3}", Button 4 <- "EMP IDB_stations_me{13}_partNumbers{4}", Button 5 <- "EMP IDB_stations_me{13}_partNumbers{5}", Button 6 <- "EMP IDB_stations_me{13}_partNumbers{6}", Button 7 <- "EMP IDB_stations_me{13}_partNumbers{7}"

recipe "CHM 04": Button 0 <- "EMP IDB_stations_me{14}_partNumbers{0}", Button 1 <- "EMP IDB_stations_me{14}_partNumbers{1}", Button 2 <- "EMP IDB_stations_me{14}_partNumbers{2}", Button 3 <- "EMP IDB_stations_me{14}_partNumbers{3}", Button 4 <- "EMP IDB_stations_me{14}_partNumbers{4}", Button 5 <- "EMP IDB_stations_me{14}_partNumbers{5}", Button 6 <- "EMP IDB_stations_me{14}_partNumbers{6}", Button 7 <- "EMP IDB_stations_me{14}_partNumbers{7}"

recipe "CHM 05": Button 0 <- "EMP IDB_stations_me{15}_partNumbers{0}", Button 1 <- "EMP IDB_stations_me{15}_partNumbers{1}", Button 2 <- "EMP IDB_stations_me{15}_partNumbers{2}", Button 3 <- "EMP IDB_stations_me{15}_partNumbers{3}", Button 4 <- "EMP IDB_stations_me{15}_partNumbers{4}", Button 5 <- "EMP IDB_stations_me{15}_partNumbers{5}", Button 6 <- "EMP IDB_stations_me{15}_partNumbers{6}", Button 7 <- "EMP IDB_stations_me{15}_partNumbers{7}"

recipe "CDO 01": Button 0 <- "EMP IDB_stations_me{16}_partNumbers{0}", Button 1 <- "EMP IDB_stations_me{16}_partNumbers{1}", Button 2 <- "EMP IDB_stations_me{16}_partNumbers{2}", Button 3 <- "EMP IDB_stations_me{16}_partNumbers{3}", Button 4 <- "EMP IDB_stations_me{16}_partNumbers{4}", Button 5 <- "EMP IDB_stations_me{16}_partNumbers{5}", Button 6 <- "EMP IDB_stations_me{16}_partNumbers{6}", Button 7 <- "EMP IDB_stations_me{16}_partNumbers{7}"

recipe "CDO 02": Button 0 <- "EMP IDB_stations_me{17}_partNumbers{0}", Button 1 <- "EMP IDB_stations_me{17}_partNumbers{1}", Button 2 <- "EMP IDB_stations_me{17}_partNumbers{2}", Button 3 <- "EMP IDB_stations_me{17}_partNumbers{3}", Button 4 <- "EMP IDB_stations_me{17}_partNumbers{4}", Button 5 <- "EMP IDB_stations_me{17}_partNumbers{5}", Button 6 <- "EMP IDB_stations_me{17}_partNumbers{6}", Button 7 <- "EMP IDB_stations_me{17}_partNumbers{7}"

recipe "CDO 03": Button 0 <- "EMP IDB_stations_me{18}_partNumbers{0}", Button 1 <- "EMP IDB_stations_me{18}_partNumbers{1}", Button 2 <- "EMP IDB_stations_me{18}_partNumbers{2}", Button 3 <- "EMP IDB_stations_me{18}_partNumbers{3}", Button 4 <- "EMP IDB_stations_me{18}_partNumbers{4}", Button 5 <- "EMP IDB_stations_me{18}_partNumbers{5}", Button 6 <- "EMP IDB_stations_me{18}_partNumbers{6}", Button 7 <- "EMP IDB_stations_me{18}_partNumbers{7}"

recipe "BFL 01": Button 0 <- "EMP IDB_stations_me{19}_partNumbers{0}", Button 1 <- "EMP IDB_stations_me{19}_partNumbers{1}", Button 2 <- "EMP IDB_stations_me{19}_partNumbers{2}", Button 3 <- "EMP IDB_stations_me{19}_partNumbers{3}", Button 4 <- "EMP IDB_stations_me{19}_partNumbers{4}", Button 5 <- "EMP IDB_stations_me{19}_partNumbers{5}", Button 6 <- "EMP IDB_stations_me{19}_partNumbers{6}", Button 7 <- "EMP IDB_stations_me{19}_partNumbers{7}"

recipe "BFL 02": Button 0 <- "EMP IDB_stations_me{20}_partNumbers{0}", Button 1 <- "EMP IDB_stations_me{20}_partNumbers{1}", Button 2 <- "EMP IDB_stations_me{20}_partNumbers{2}", Button 3 <- "EMP IDB_stations_me{20}_partNumbers{3}", Button 4 <- "EMP IDB_stations_me{20}_partNumbers{4}", Button 5 <- "EMP IDB_stations_me{20}_partNumbers{5}", Button 6 <- "EMP IDB_stations_me{20}_partNumbers{6}", Button 7 <- "EMP IDB_stations_me{20}_partNumbers{7}"

recipe "BFL 03": Button 0 <- "EMP IDB_stations_me{21}_partNumbers{0}", Button 1 <- "EMP IDB_stations_me{21}_partNumbers{1}", Button 2 <- "EMP IDB_stations_me{21}_partNumbers{2}", Button 3 <- "EMP IDB_stations_me{21}_partNumbers{3}", Button 4 <- "EMP IDB_stations_me{21}_partNumbers{4}", Button 5 <- "EMP IDB_stations_me{21}_partNumbers{5}", Button 6 <- "EMP IDB_stations_me{21}_partNumbers{6}", Button 7 <- "EMP IDB_stations_me{21}_partNumbers{7}"

recipe "LGS 01": Button 0 <- "EMP IDB_stations_me{22}_partNumbers{0}", Button 1 <- "EMP IDB_stations_me{22}_partNumbers{1}", Button 2 <- "EMP IDB_stations_me{22}_partNumbers{2}", Button 3 <- "EMP IDB_stations_me{22}_partNumbers{3}", Button 4 <- "EMP IDB_stations_me{22}_partNumbers{4}", Button 5 <- "EMP IDB_stations_me{22}_partNumbers{5}", Button 6 <- "EMP IDB_stations_me{22}_partNumbers{6}", Button 7 <- "EMP IDB_stations_me{22}_partNumbers{7}"

recipe "LGS 02": Button 0 <- "EMP IDB_stations_me{23}_partNumbers{0}", Button 1 <- "EMP IDB_stations_me{23}_partNumbers{1}", Button 2 <- "EMP IDB_stations_me{23}_partNumbers{2}", Button 3 <- "EMP IDB_stations_me{23}_partNumbers{3}", Button 4 <- "EMP IDB_stations_me{23}_partNumbers{4}", Button 5 <- "EMP IDB_stations_me{23}_partNumbers{5}", Button 6 <- "EMP IDB_stations_me{23}_partNumbers{6}", Button 7 <- "EMP IDB_stations_me{23}_partNumbers{7}"

screen "1 PART CALL" 1366x768
   on GenerateScreen: SetTag("HMI_screenNumber", 1)
   Rectangle "Settings Tab Background" at 682,0 size 684x68
      Appearance <- "HMI_screenNumber"
   Rectangle "Part Call Tab Background" at 0,0 size 685x68
      Appearance <- "HMI_screenNumber"
   Rectangle "Settings Tab Border Hide" at 685,61 size 678x20
      Visibility <- "HMI_screenNumber"
   Rectangle "Part Call Tab Border Hide" at 3,61 size 679x20
      Visibility <- "HMI_screenNumber"
   Button "Settings Screen" at 683,0 size 683x68; TextOff 'SETTINGS'; Authorization "User administration"
      on Release: ActivateScreen("2 SETTINGS", 0)
   Button "Part Call Screen" at 0,0 size 683x68; TextOff 'PART CALL'
      on Release: ActivateScreen("1 PART CALL", 0)
   TextField "Header Line" at 32,112 size 216x53; Text 'LINE'
   TextField "Header Drop Zone" at 238,112 size 236x53; Text 'DROP ZONE'
   TextField "Header Part Number" at 474,112 size 648x53; Text 'PART NUMBER'
   TextField "Header Time" at 1112,112 size 222x53; Text 'TIME'
   ScreenModuleView "TableRow00" at 27,170 size 1312x52; ScreenModuleType ""
      Guid_{11997190-27688} <- "HMI_partCall_row{0}"
      on Guid_{11997190-83214}: ActivateScreen("3 BARCODE", 0)
   ScreenModuleView "TableRow01" at 27,222 size 1312x52; ScreenModuleType ""
      Guid_{11997190-27688} <- "HMI_partCall_row{1}"
      on Guid_{11997190-83214}: ActivateScreen("3 BARCODE", 0)
   ScreenModuleView "TableRow02" at 27,274 size 1312x52; ScreenModuleType ""
      Guid_{11997190-27688} <- "HMI_partCall_row{2}"
      on Guid_{11997190-83214}: ActivateScreen("3 BARCODE", 0)
   ScreenModuleView "TableRow03" at 27,326 size 1312x52; ScreenModuleType ""
      Guid_{11997190-27688} <- "HMI_partCall_row{3}"
      on Guid_{11997190-83214}: ActivateScreen("3 BARCODE", 0)
   ScreenModuleView "TableRow04" at 27,378 size 1312x52; ScreenModuleType ""
      Guid_{11997190-27688} <- "HMI_partCall_row{4}"
      on Guid_{11997190-83214}: ActivateScreen("3 BARCODE", 0)
   ScreenModuleView "TableRow05" at 27,430 size 1312x52; ScreenModuleType ""
      Guid_{11997190-27688} <- "HMI_partCall_row{5}"
      on Guid_{11997190-83214}: ActivateScreen("3 BARCODE", 0)
   ScreenModuleView "TableRow06" at 27,482 size 1312x52; ScreenModuleType ""
      Guid_{11997190-27688} <- "HMI_partCall_row{6}"
      on Guid_{11997190-83214}: ActivateScreen("3 BARCODE", 0)
   ScreenModuleView "TableRow07" at 27,534 size 1312x52; ScreenModuleType ""
      Guid_{11997190-27688} <- "HMI_partCall_row{7}"
      on Guid_{11997190-83214}: ActivateScreen("3 BARCODE", 0)
   ScreenModuleView "TableRow08" at 27,586 size 1312x52; ScreenModuleType ""
      Guid_{11997190-27688} <- "HMI_partCall_row{8}"
      on Guid_{11997190-83214}: ActivateScreen("3 BARCODE", 0)
   ScreenModuleView "TableRow09" at 27,638 size 1312x52; ScreenModuleType ""
      Guid_{11997190-27688} <- "HMI_partCall_row{9}"
      on Guid_{11997190-83214}: ActivateScreen("3 BARCODE", 0)
   ScreenModuleView "TableRow10" at 27,690 size 1312x52; ScreenModuleType ""
      Guid_{11997190-27688} <- "HMI_partCall_row{10}"
      on Guid_{11997190-83214}: ActivateScreen("3 BARCODE", 0)

